   // Kleine Einschatverzögerung
         L     #Temp_SetValueTemp;
         L     "DB751_auxiliaryDriveMetering".HeatexchangerLP[1].Offset_Cooling;
         +R;
         L     #Temp_ND_WT;
         >R;
         =     #Temp_MoreDelta;
   // Kühlen  AUS
         L     "DB613_Komponent_State".HeatexchangerLP[1].PulsTime;
         RND;
         L     #Zeit_abgelaufen;
         <D;
         AN(;
         L     "DB613_Komponent_State".HeatexchangerLP[1].PulsTime;
         RND;
         L     #Regelstrecke;
         >D;
         );
         ON    "DB613_Komponent_State".HeatexchangerLP[1].Switch_Temp_ON_OFF;
         ON    "DB619_State_MPart".Operationmode[1].valid;
         O     "DB823_Error_Metering".Temperature_HeatexchangerLP[1].Sensor_FLT_broken_wire;
         O     #Temp_MoreDelta;
         R     "DB613_Komponent_State".HeatexchangerLP[1].CoolingActive;

   // Valve in FB101 for Heatexchanger in back run
   //      =     "V_Heatexchanger_C1" // stromlos zu

   //-----
   // Check limits temperature 1 Heatexchanger

         CALL  "FC916_PV_Limits"
         ( IN_Tolerance_Test     := "DB619_State_MPart".Operationmode[1].Controllvoltage,
           IN_Reset_Fault        := "DB009_Faults".Faults_Reset_FKT_M1,
           IO_Any_ArrayPV        := "DB608_PV_Metering".HeatexchangerLP[1],
           IO_Fault_Warn_upperL  := "DB823_Error_Metering".Temperature_HeatexchangerLP[1].Warning_limit_plus,
           IO_Fault_Warn_lowerL  := "DB823_Error_Metering".Temperature_HeatexchangerLP[1].Warning_limit_minus,
           IO_Fault_Alarm_upperL := "DB823_Error_Metering".Temperature_HeatexchangerLP[1].Alarm_limit_plus,
           IO_Fault_Alarm_lowerL := "DB823_Error_Metering".Temperature_HeatexchangerLP[1].Alarm_limit_minus,
           IO_New_Fault          := "DB009_Faults".Faultschanging_M1,
           IO_Fault_Level_1      := "DB009_Faults".Faults_FKT_Grp_1_M1,
           IO_Fault_Level_2      := "DB009_Faults".Faults_FKT_Grp_2_M1,
           IO_Fault_Level_3      := "DB009_Faults".Faults_FKT_Grp_3_M1
         );
   //-----
   // State of Switch
         L     0;
         A     "DB613_Komponent_State".HeatexchangerLP[1].CoolingActive;
         A     "DB619_State_MPart".Machine[1].Metering."01";
         A     "DB613_Komponent_State".HeatexchangerLP[1].Switch_Temp_ON_OFF;
         JCN   S1H1;
         L     1;
   S1H1: ON    "DB613_Komponent_State".HeatexchangerLP[1].CoolingActive;
         ON    "DB619_State_MPart".Machine[1].Metering."01";
         A     "DB613_Komponent_State".HeatexchangerLP[1].Switch_Temp_ON_OFF;
         JCN   S2H1;
         L     3;
   S2H1: A     "DB823_Error_Metering".Temperature_HeatexchangerLP[1].Sensor_FLT_broken_wire;
         A     "DB613_Komponent_State".HeatexchangerLP[1].Switch_Temp_ON_OFF;
         JCN   S3H1;
         L     2;
   S3H1: T     "DB613_Komponent_State".HeatexchangerLP[1].State_Temp;
   EHD1: NOP   0;

   // Fault exists
         O     "DB823_Error_Metering".Temperature_HeatexchangerLP[1].Sensor_FLT_broken_wire;
         O     "DB823_Error_Metering".Temperature_HeatexchangerLP[1].Warning_limit_plus;
         O     "DB823_Error_Metering".Temperature_HeatexchangerLP[1].Warning_limit_minus;
         O     "DB823_Error_Metering".Temperature_HeatexchangerLP[1].Alarm_limit_plus;
         O     "DB823_Error_Metering".Temperature_HeatexchangerLP[1].Alarm_limit_minus;
         =     "DB613_Komponent_State".HeatexchangerLP[1].Fault_Exist;
END_REGION

REGION Network 2: There is no connection to the sensor (3)
   //---------------------------------------------
   //  Controller temperature Heatexchanger K2
   //---------------------------------------------
         AN    "DB753_MeteringPump".Pump[2].WithLPHeatExchanger;
         R     "DB823_Error_Metering".Temperature_HeatexchangerLP[2].Sensor_FLT_broken_wire;
         R     "DB823_Error_Metering".Temperature_HeatexchangerLP[2].Warning_limit_plus;
         R     "DB823_Error_Metering".Temperature_HeatexchangerLP[2].Warning_limit_minus;
         R     "DB823_Error_Metering".Temperature_HeatexchangerLP[2].Alarm_limit_plus;
         R     "DB823_Error_Metering".Temperature_HeatexchangerLP[2].Alarm_limit_minus;
         R     "DB613_Komponent_State".HeatexchangerLP[2].Fault_Exist;
         JC    EHD2;
   //-----
         CALL  "FC920_PV_Calc_Act_Value"
         ( IN_Act_Value_read := TRUE,
           IN_Act_Value_ext  := FALSE,
           IN_Ext_Value      := #DINT_dummy,
           IN_Read_Double    := FALSE,
           IN_FLT_Needful    := 1,
           IN_FLT_Reset      := "DB009_Faults".Faults_Reset_FKT_M1,
           IO_Any_ArrayPV    := "DB608_PV_Metering".HeatexchangerLP[2],
           IO_Fault_Sensor   := "DB823_Error_Metering".Temperature_HeatexchangerLP[2].Sensor_FLT_broken_wire,
           IO_New_Fault      := "DB009_Faults".Faultschanging_M1,
           IO_FLT_Level_3    := "DB009_Faults".Faults_FKT_Grp_3_M1
         );
   //
         L     "DB608_PV_Metering".HeatexchangerLP[2].PV_ActV.Value;
         DTR;
         L     10.0;
         /R;
         T     #Temp_ND_WT;
   //
         L     "DB608_PV_Metering".HeatexchangerLP[2].PV_SetV.Value;
         DTR;
         L     10.0;
         /R;
         T     #Temp_SetValueTemp;
   //
         CALL  "FC056_TemPulse2"
         ( Trig              := "Start_Controler1_LP_K2",
           In_Sollwert       := #Temp_SetValueTemp,
           In_Istwert_Tank   := #Temp_ND_WT,
           In_Istwert_Return := #Temp_ND_WT,
           In_Wichtung       := "DB751_auxiliaryDriveMetering".HeatexchangerLP[2].Weighting_Temp,
           In_Regelstrecke   := "DB751_auxiliaryDriveMetering".HeatexchangerLP[2].PLC_Control_Area,
           In_MaxDelta_K     := "DB751_auxiliaryDriveMetering".HeatexchangerLP[2].Max_Temp_Diff_Cooling,
           In_MaxDelta_H     := "DB751_auxiliaryDriveMetering".HeatexchangerLP[2].Max_Temp_Diff_Heating,
           Pulsezeit         := "DB613_Komponent_State".HeatexchangerLP[2].PulsTime,
           Heating           := #Dummy,
           Cooling           := #Temp_Cooling
         );
   //
   //Regelstrecke ms Format
         L     "DB751_auxiliaryDriveMetering".HeatexchangerLP[2].PLC_Control_Area;
         L     1000.0;
         *R;
         RND;
         T     #Regelstrecke;  // Zeitwert für Timer

   // Regelstreckentimer ständig starten

         AN    "Start_Controler1_LP_K2";
         =     "Start_Controler2_LP_K2";

         CALL  TON , "DB61_Temp_ND_WT_MK1_K2"
         ( IN := "Start_Controler2_LP_K2",
           PT := #Regelstrecke,
           Q  := "Start_Controler1_LP_K2",
           ET := #Zeit_abgelaufen
         );

   // Kühlen  EIN
         A     #Temp_Cooling;
         S     "DB613_Komponent_State".HeatexchangerLP[2].CoolingActive;

   //Kleine Einschatverzögerung
         L     #Temp_SetValueTemp;
         L     "DB751_auxiliaryDriveMetering".HeatexchangerLP[2].Offset_Cooling;
         +R;
         L     #Temp_ND_WT;
         >R;
         =     #Temp_MoreDelta;

   // Kühlen  AUS
         L     "DB613_Komponent_State".HeatexchangerLP[2].PulsTime;
         RND;
         L     #Zeit_abgelaufen;
         <D;
         AN(;
         L     "DB613_Komponent_State".HeatexchangerLP[2].PulsTime;
         RND;
         L     #Regelstrecke;
         >D;
         );
         ON    "DB613_Komponent_State".HeatexchangerLP[2].Switch_Temp_ON_OFF;
         ON    "DB619_State_MPart".Operationmode[1].valid;
         O     "DB823_Error_Metering".Temperature_HeatexchangerLP[2].Sensor_FLT_broken_wire;
         O     #Temp_MoreDelta;
         R     "DB613_Komponent_State".HeatexchangerLP[2].CoolingActive;

   // Valve in FB102 for Heatexchanger in back run
   //     =     "V_Heatexchanger_C2" // stromlos zu


   //-----
   // Check limits temperature 2 Heatexchanger

         CALL  "FC916_PV_Limits"
         ( IN_Tolerance_Test     := "DB619_State_MPart".Operationmode[1].Controllvoltage,
           IN_Reset_Fault        := "DB009_Faults".Faults_Reset_FKT_M1,
           IO_Any_ArrayPV        := "DB608_PV_Metering".HeatexchangerLP[2],
           IO_Fault_Warn_upperL  := "DB823_Error_Metering".Temperature_HeatexchangerLP[2].Warning_limit_plus,
           IO_Fault_Warn_lowerL  := "DB823_Error_Metering".Temperature_HeatexchangerLP[2].Warning_limit_minus,
           IO_Fault_Alarm_upperL := "DB823_Error_Metering".Temperature_HeatexchangerLP[2].Alarm_limit_plus,
           IO_Fault_Alarm_lowerL := "DB823_Error_Metering".Temperature_HeatexchangerLP[2].Alarm_limit_minus,
           IO_New_Fault          := "DB009_Faults".Faultschanging_M1,
           IO_Fault_Level_1      := "DB009_Faults".Faults_FKT_Grp_1_M1,
           IO_Fault_Level_2      := "DB009_Faults".Faults_FKT_Grp_2_M1,
           IO_Fault_Level_3      := "DB009_Faults".Faults_FKT_Grp_3_M1
         );
   //-----
   // State of Switch
         L     0;
         A     "DB613_Komponent_State".HeatexchangerLP[2].CoolingActive;
         A     "DB619_State_MPart".Machine[1].Metering."02";
         A     "DB613_Komponent_State".HeatexchangerLP[2].Switch_Temp_ON_OFF;
         JCN   S1H2;
         L     1;
   S1H2: ON    "DB613_Komponent_State".HeatexchangerLP[2].CoolingActive;
         ON    "DB619_State_MPart".Machine[1].Metering."02";
         A     "DB613_Komponent_State".HeatexchangerLP[2].Switch_Temp_ON_OFF;
         JCN   S2H2;
         L     3;
   S2H2: A     "DB823_Error_Metering".Temperature_HeatexchangerLP[2].Sensor_FLT_broken_wire;
         A     "DB613_Komponent_State".HeatexchangerLP[2].Switch_Temp_ON_OFF;
         JCN   S3H2;
         L     2;
   S3H2: T     "DB613_Komponent_State".HeatexchangerLP[2].State_Temp;
   EHD2: NOP   0;

   // Fault exists
         O     "DB823_Error_Metering".Temperature_HeatexchangerLP[2].Sensor_FLT_broken_wire;
         O     "DB823_Error_Metering".Temperature_HeatexchangerLP[2].Warning_limit_plus;
         O     "DB823_Error_Metering".Temperature_HeatexchangerLP[2].Warning_limit_minus;
         O     "DB823_Error_Metering".Temperature_HeatexchangerLP[2].Alarm_limit_plus;
         O     "DB823_Error_Metering".Temperature_HeatexchangerLP[2].Alarm_limit_minus;
         =     "DB613_Komponent_State".HeatexchangerLP[2].Fault_Exist;
END_REGION
END_FUNCTION

FUNCTION "FC071_CleaningPiston" : Void   // FC71, STL
TITLE = Function of cleaning piston mixing head
{ S7_Optimized_Access := 'FALSE' }
AUTHOR : KT242
FAMILY : RS_KK
NAME : CP
VERSION : 1.3
   VAR_INPUT
      IN_WithCP : Bool;   // Signal cleaning piston exists at mixinghead
      IN_Ana_CP_State : Byte;   // State of analog cleaning piston
      IN_SWUEnabled : Bool;   // Switch over unit for this mixing head is enabled
      IN_ButtonCPForward : Bool;   // Button cleaning piston manually forward
      IN_ButtonCPback : Bool;   // Button cleaning piston manually back
      IN_CPForwardFromExternal : Bool;   // External signal (e.g. from robot) to move the CP forward
      IN_CPAfterShot : Bool;   // Signal cleaning piston has to move after the shot
      IN_PartshotDisabled : Bool;   // Partshot disabled -> like service shot
      IN_Blowing_OUT : Bool;   // Blowing out after Shot
      IN_CPProxSwitch : Bool;   // Proximity switch cleaning piston is back (rest position)
      IN_SWUActive : Bool;   // Only this switch over unit is activated
      IN_HydraulicOk : Bool;   // Hydraulic ok
      IN_ResetFaults : Bool;   // Signal to reset error bits
      IN_ControlVoltage : Bool;   // Control Voltage is on
      IN_OperatingModeValid : Bool;   // Valid operating mode is activated
      IN_OperatingModeWithFoam : Bool;   // Machine is not in service mode (this is a condition for cleaning)
      IN_OperatingModeTestValv : Bool;   // Machine is in mode test with test valves (no cleaning necessary)
      IN_Lamptest : Bool;   // Lamptest selected
      IN_ShotEnd : Bool;   // Ramp shot finished
      IN_FaultLevel_1 : Bool;   // Fault level 1 on machine
      IN_PressurizeTimeRunning : Bool;   // Time for building up pressure and flow values is active
      IN_ShotActive : Bool;   // Shot is active
      IN_CycleRunning : Bool;   // Shotcycle is active
      IN_RmpCtrlChangeTimeEnd : Bool;   // Recirculation between shots finished
      IN_StandbyTimeRunning : Bool;   // Recirculation after shot acvtiv
      IN_RmpCycleEnd : Bool;   // Foaming cycle finished
      IN_CPTimer : Timer;   // Timer for CP-funkctions
      IN_TMCheckHomePos : Timer;   // Timer to suppress fault homepos when module begins regulation
      Values : "UDT771_CleaningPiston";
   END_VAR
   VAR_IN_OUT
      OUT_ValveCPForward : Bool;   // Valve to move the CP forward
      OUT_LampCPBack : Bool;   // Lamp to display that the CP is back
      IO_CPIsOk : Bool;   // CP is ok -> enables shot
      IO_ReqHydrForCleaning : Bool;   // Request hydraulic pressure for cleaning stroke
      IO_Status : ANY;   // Status flags for CP
      IO_Fault : ANY;
      IO_NewFault : Bool;
      IO_FaultLevel_1 : Bool;
      IO_FaultLevel_2 : Bool;
      IO_FaultLevel_3 : Bool;
   END_VAR
   VAR_TEMP
      Temp_IO_Status : "UDT071_CPiston_State";
      TEMP_IO_Fault : "UDT1871_FLT_CPiston";
      ERROR_CODE : Int;   // Error state of systemfunction "BLKMOV" Blockmove
      Anypointer1 : ANY;   // Pointer to copy thr array "IO_Status" and "Temp_IO_Status"
      Anypointer2 : ANY;   // Pointer to copy thr array "IO_Status" and "Temp_IO_Status"
      InterruptCleaningStroke : Bool;   // Flag of interrupt cleaning cycle
      StartCleaningStroke : Bool;   // Flag cleaning cycle started
      ShotFinished : Bool;   // Flag activate cleaning piston after part shot
      TempAnaCPBack : Bool;   // Analog controlled leaning piston is back
      WrongType : Bool;   // Wrong Mixing Head Type
   END_VAR
BEGIN

REGION Network 1: Saved data integration
         LAR1;
         L;
         LAR2;
   //
         L     16#1002;  // Bytes
         T     W[AR1, P#0.0];
         L     W[AR2, P#2.0];  // Amount of bytes
         T     W[AR1, P#2.0];
         L     W[AR2, P#4.0];  // Block no,
         T     W[AR1, P#4.0];
         L     D[AR2, P#6.0];  // Startadress of datas
         T     D[AR1, P#6.0];
   //
         CALL  BLKMOV
         ( SRCBLK  := #Anypointer1,
           RET_VAL := #ERROR_CODE,
           DSTBLK  := #Temp_IO_Status
         );
   //
         LAR1;
         L;
         LAR2;
   //
         L     16#1002;  // Bytes
         T     W[AR1, P#0.0];
         L     W[AR2, P#2.0];  // Amount of bytes
         T     W[AR1, P#2.0];
         L     W[AR2, P#4.0];  // Block no,
         T     W[AR1, P#4.0];
         L     D[AR2, P#6.0];  // Startadress of datas
         T     D[AR1, P#6.0];
   //
         CALL  BLKMOV
         ( SRCBLK  := #Anypointer2,
           RET_VAL := #ERROR_CODE,
           DSTBLK  := #TEMP_IO_Fault
         );
   //
         A(;
         L     #IN_Ana_CP_State;
         AW    16#0080;
         A     <>0;
         );
         A(;
         O     #Values.ContrCleaningPiston;
         O     #Values.StepCleaningPiston;
         );
         =     #TempAnaCPBack;
END_REGION

REGION Network 2: Cleaning stroke forward
         AN    #IN_WithCP;
         R     #Values.Spare_19;

         ON    #IN_WithCP;
         ON    #Values.Spare_19;
         R     #Temp_IO_Status.Switch_CP_Forward;

         NOT;
         CLR;
         =     #WrongType;
         A     #WrongType;
         JC    STG;
END_REGION

REGION Network 3: CP existing or not?
         O     #IN_CPProxSwitch;
         O     #TempAnaCPBack;
         AN    #TEMP_IO_Fault.IPS_defect;
         ON    #IN_WithCP;
         A     #IN_SWUActive;
         =     #Temp_IO_Status.CP_is_OK;
         S     #IO_CPIsOk;
   //
         A     #Temp_IO_Status.CP_is_OK;
         FN    #Temp_IO_Status.Edge_CP_nOK;
         R     #IO_CPIsOk;
   //
         A     #IN_SWUEnabled;
         A     #IN_WithCP;
         JC    STG;
   //
         SET;
         R     #Temp_IO_Status.MH_was_open;
         R     #Temp_IO_Status.Cleaning_runs;
         R     #Temp_IO_Status.CleaningFromEPrunning;
         R     #Temp_IO_Status.CleanAfterShotSelected;
         R     #Temp_IO_Status.Stop_Cleaning;
         R     #Temp_IO_Status.CP_valve_selected;
         R     #Temp_IO_Status.CP_Moved_Manual;
         R     #Temp_IO_Status.FaultExists;
         R     #TEMP_IO_Fault.Forward_to_slow;
         R     #TEMP_IO_Fault.Back_to_slow;
         R     #TEMP_IO_Fault.IPS_defect;
         R     #TEMP_IO_Fault.Lost_IPS_position;
         L     0;
         T     #Temp_IO_Status.Stepnumber;
   //
         JU    LAMP;
END_REGION

REGION Network 4: Error handling
   STG:  NOP   0;
   // Reset faults
         A     #IN_ResetFaults;
         R     #TEMP_IO_Fault.Lost_IPS_position;
         R     #TEMP_IO_Fault.IPS_defect;
         R     #TEMP_IO_Fault.Forward_to_slow;
         R     #TEMP_IO_Fault.Back_to_slow;
         R     #TEMP_IO_Fault.Leaves_HomePos;
   //
         A     #WrongType;
         JC    err;

   // Fault No.1: Cleaning piston leaves the backward position during shot
         L     2#0000_0000_0000_0100;
         L     #IN_Ana_CP_State;
         AW;
         L     0;
         >D;
         A(;
         O     #Values.ContrCleaningPiston;
         O     #Values.StepCleaningPiston;
         );
         O;
         A     #IN_SWUActive;
         A     #IN_ShotActive;
         AN(;
         O     #Values.ContrCleaningPiston;
         O     #Values.StepCleaningPiston;
         );
         AN    #IN_CPProxSwitch;
         AN    #TEMP_IO_Fault.Lost_IPS_position;
         S     #TEMP_IO_Fault.Lost_IPS_position;
         S     #IO_NewFault;
   //
   // Fault No.2: Priximity switch cleaning piston back is broken
         AN    #IN_CPProxSwitch;
         A     #IN_HydraulicOk;
         AN    #TEMP_IO_Fault.Back_to_slow;
         AN    #Temp_IO_Status.Cleaning_runs;
         AN(;
         O     #Values.ContrCleaningPiston;
         O     #Values.StepCleaningPiston;
         );
         AN    #TEMP_IO_Fault.Lost_IPS_position;
         AN    #TEMP_IO_Fault.IPS_defect;
         S     #TEMP_IO_Fault.IPS_defect;
         S     #IO_NewFault;
   //
   // Fault No. 3: Movement forward of analog cleaning piston too slow
         L     2#0000_0000_0000_0001;
         L     #IN_Ana_CP_State;
         AW;
         L     0;
         >D;
         A(;
         O     #Values.ContrCleaningPiston;
         O     #Values.StepCleaningPiston;
         );
         AN    #TEMP_IO_Fault.Forward_to_slow;
         S     #TEMP_IO_Fault.Forward_to_slow;
         S     #IO_NewFault;
   // Fault No. 3: Movement forward of cleaning piston too slow is build later
   //

   // Fault No. 4: Movement back of analog cleaning piston too slow
         L     2#0000_0000_0000_0010;
         L     #IN_Ana_CP_State;
         AW;
         L     0;
         >D;
         A(;
         O     #Values.ContrCleaningPiston;
         O     #Values.StepCleaningPiston;
         );
         AN    #TEMP_IO_Fault.Back_to_slow;
         S     #TEMP_IO_Fault.Back_to_slow;
         S     #IO_NewFault;
   // Fault No. 4: Movement back of cleaning piston too slow is build later
   //
   // Fault No. 14: Cleaning piston is leaving home position
   //
         A     #IN_HydraulicOk;
         L     S5T#500MS;
         SD    #IN_TMCheckHomePos;
         A(;
         L     2#0000_0000_0010_0000;
         L     #IN_Ana_CP_State;
         AW;
         L     0;
         >D;
         );
         A(;
         O     #Values.ContrCleaningPiston;
         O     #Values.StepCleaningPiston;
         );
         A     #IN_TMCheckHomePos;
         AN    #TEMP_IO_Fault.Leaves_HomePos;
         S     #TEMP_IO_Fault.Leaves_HomePos;
         S     #IO_NewFault;
END_REGION

REGION Network 5: Error handling
   err:  NOP   0;
         O     #TEMP_IO_Fault.Forward_to_slow;
         O     #TEMP_IO_Fault.Back_to_slow;
         O     #TEMP_IO_Fault.IPS_defect;
         O     #TEMP_IO_Fault.Lost_IPS_position;
         O     #TEMP_IO_Fault.Leaves_HomePos;
         =     #Temp_IO_Status.FaultLevel_1;
         =     #Temp_IO_Status.FaultExists;
         S     #IO_FaultLevel_1;

         CLR;
         =     #Temp_IO_Status.FaultLevel_2;
         S     #IO_FaultLevel_2;

         CLR;
         =     #Temp_IO_Status.FaultLevel_3;
         S     #IO_FaultLevel_3;

         A     #WrongType;
         JC    LAMP;
END_REGION

REGION Network 6: Cleaning necessary or not
   // Step 1: Detect if the mixinghead was open.
   //         The signal is built newly for each partshot and only if the mixinghead
   //         was really opened a cleaning stroke is carried out
   //         -> "Temp_IO_Status.MH_was_open"
   //         It is reset when:
   //         - the switching unit is deselected
   //         - a new shot is started (no matter on wich mixinghead)
   //         - the shot cycle is finished
   //         - the cleaning stroke was done
   //         - the operating mode is deselected
   // 
   // Step 2: If for this shot a cleaning stroke was selected or after fault group 1
   //         the cleaning piston moves forward.
   //         -> "Temp_IO_Status.Cleaning_a_Shot_selected"
   //         The bit is reset if:
   //         - the switching unit is deselected
   //         - the cleaning stroke was done 
   //         - the operating mode is deselected
         A     #IN_ShotActive;
         A     #IN_OperatingModeWithFoam;
         AN    #IN_PartshotDisabled;
         AN    #IN_OperatingModeTestValv;
         A     #IN_SWUActive;
         S     #Temp_IO_Status.MH_was_open;
   //
         A     #IN_CPAfterShot;
         A     #IN_ShotEnd;
         O     #IN_FaultLevel_1;
         ON    #IN_ControlVoltage;
         A     #Temp_IO_Status.MH_was_open;
         S     #Temp_IO_Status.CleanAfterShotSelected;
   //
         O     #Temp_IO_Status.CleanAfterShotSelected;
         O     #IN_RmpCtrlChangeTimeEnd;
         O     #Temp_IO_Status.Stop_Cleaning;
         ON    #IN_OperatingModeValid;
         R     #Temp_IO_Status.MH_was_open;
   //
END_REGION

REGION Network 7: Interrupt cleaning stroke
   // A cleaning cycle is interrupted in the following cases:
   //            - Button cleaning piston back is used without acting the butten
   //              cleaning piston forward at the same time  (LFI) 
   //            - The robot resets the signal cleaning piston forward
   //            - a new shot is being started on this mixinghead
   // 
   // If a cleaning stroke should be interrupted, the step counter for the cleaning
   // cycle is set to 6 (reset output for valve CP forward)
         A(;
         O     #IN_PressurizeTimeRunning;
         O     #IN_RmpCtrlChangeTimeEnd;
         A     #IN_SWUActive;
         O;
         A     #Temp_IO_Status.CleaningFromEPrunning;
         AN    #IN_CPForwardFromExternal;
         O;
         A     #IN_ButtonCPback;
         );
         A     #Temp_IO_Status.Cleaning_runs;
         AN    #Temp_IO_Status.Stop_Cleaning;
         S     #Temp_IO_Status.Stop_Cleaning;
         =     #InterruptCleaningStroke;
   //
         AN    #InterruptCleaningStroke;
         JC    CONT;
   //
         L     6;
         T     #Temp_IO_Status.Stepnumber;
   //
   CONT: A     #IN_CPForwardFromExternal;
         =     #Temp_IO_Status.CleaningFromEPrunning;
END_REGION

REGION Network 8: Start cleaning stroke
   //  1. Block:
   //
         A(;
   // A.:
         O     #IN_ButtonCPForward;
         O     #Temp_IO_Status.Switch_CP_Forward;
         AN    #IN_ButtonCPback;
         O     #Temp_IO_Status.CleaningFromEPrunning;
         A(;
         ON    #IN_CycleRunning;
         O     #IN_StandbyTimeRunning;
         ON    #IN_SWUActive;
         );
   // B.:
         O(;
         A     #IN_ShotEnd;
         A     #Temp_IO_Status.CleanAfterShotSelected;
         );
         );
         A     #IN_HydraulicOk;
   //  2. Block:
   //
         O(;
         ON    #IN_ControlVoltage;
         O     #IN_FaultLevel_1;
         A     #Temp_IO_Status.CleanAfterShotSelected;
         );
   // für alle:
         AN    #Temp_IO_Status.Stop_Cleaning;
         AN    #Temp_IO_Status.Cleaning_runs;
         S     #Temp_IO_Status.Cleaning_runs;
         =     #StartCleaningStroke;
   //
         AN    #StartCleaningStroke;
         JC    STEP;
   //
         A     #IN_ButtonCPForward;
         S     #Temp_IO_Status.CP_Moved_Manual;
         L     1;
         T     #Temp_IO_Status.Stepnumber;
   STEP: NOP   0;
END_REGION

REGION Network 9: organize steps of cleaning stroke
         L     #Temp_IO_Status.Stepnumber;
         JL    DEL;  // if step number > 7 or
         JU    DEL;  // 0: delete
         JU    ST1;  // 1: check if waiting time back needs to be started
         JU    ST2;  // 2: start waiting time back
         JU    ST3;  // 3: actuate the valve
         JU    ST4;  // 4: monitor movement time forward
         JU    ST5;  // 5: start wait time in front
         JU    ST6;  // 6: switch off valve for CP
         JU    ST7;  // 7: monitor movement back
   //
   DEL:  CLR;  // delete status informations
         =     #Temp_IO_Status.CP_valve_selected;
         =     #Temp_IO_Status.Cleaning_runs;
         =     #Temp_IO_Status.Stop_Cleaning;
         CLR;
         SP    #IN_CPTimer;
         JU    LAMP;
END_REGION

REGION Network 10: check: wait time back necessary
   ST1:  SET;
         R     #Temp_IO_Status.Stop_Cleaning;
   //
         A     #Temp_IO_Status.CleanAfterShotSelected;
         JCN   ST1E;
         L     2;  // start waiting time back (if automatic cleaning stroke)
         T     #Temp_IO_Status.Stepnumber;
         JU    LAMP;
   //
   ST1E: L     3;  // start cleaning directly (in other cases)
         T     #Temp_IO_Status.Stepnumber;
         JU    LAMP;
END_REGION

REGION Network 11: start waiting time back
   // The waitint time back normally is 0.2 seconds
   ST2:  AN    #IN_Blowing_OUT;
         L     #Values.RestTimeBack;
         SD    #IN_CPTimer;
         AN    #IN_CPTimer;
         JC    LAMP;
   //
         L     3;
         T     #Temp_IO_Status.Stepnumber;
         CLR;
         SP    #IN_CPTimer;
         JU    LAMP;
END_REGION

REGION Network 12: Actuate the valve
   ST3:  SET;
         S     #Temp_IO_Status.CP_valve_selected;
         S     #IO_ReqHydrForCleaning;
         L     4;
         T     #Temp_IO_Status.Stepnumber;
         JU    LAMP;
END_REGION

REGION Network 13: Monitor movement time forward
   // the monitoring time is fix on 2 seconds
   ST4:  O     #IN_CPProxSwitch;  // next step when prximity switch is off
         O     #TempAnaCPBack;
         JC    LZVW;
   //
         L     5;
         T     #Temp_IO_Status.Stepnumber;
         CLR;
         SP    #IN_CPTimer;
         JU    LAMP;
   //
   LZVW: L     S5T#2S;
         SD    #IN_CPTimer;
         A     #IN_CPTimer;
         JCN   LAMP;
   //
   // Fault No.3: movement forward too slow
   //
         R     #Temp_IO_Status.CleanAfterShotSelected;
         AN    #TEMP_IO_Fault.Forward_to_slow;
         S     #TEMP_IO_Fault.Forward_to_slow;
         S     #IO_NewFault;
         L     0;
         T     #Temp_IO_Status.Stepnumber;
         JU    LAMP;
END_REGION

REGION Network 14: Wait time in fromt
   //-----
   ST5:  SET;
         R     #Temp_IO_Status.CleanAfterShotSelected;
   //-----
         A     #Temp_IO_Status.CP_Moved_Manual;
         L     #Values.RestTimeFrontManual;
         JC    TimeCPForward;
         L     #Values.RestTimeFront;
   //-----
   TimeCPForward:NOP   0;
         SET;
         SD    #IN_CPTimer;
   //-----
         A     #IN_CPTimer;
         AN    #IN_ButtonCPForward;
         AN    #Temp_IO_Status.Switch_CP_Forward;
         AN    #Temp_IO_Status.CleaningFromEPrunning;
         JCN   LAMP;
   //-----
         L     6;
         T     #Temp_IO_Status.Stepnumber;
         CLR;
         SP    #IN_CPTimer;
         JU    LAMP;
   //-----
END_REGION

REGION Network 15: switch off the valve
   ST6:  SET;
         S     #Temp_IO_Status.Stop_Cleaning;
         R     #Temp_IO_Status.CP_valve_selected;
         R     #Temp_IO_Status.CP_Moved_Manual;
         S     #IO_ReqHydrForCleaning;
         L     7;
         T     #Temp_IO_Status.Stepnumber;
         CLR;
         SP    #IN_CPTimer;
         JU    LAMP;
END_REGION

REGION Network 16: monitoring movement back
   ST7:  CLR;
         AN    #IN_CPProxSwitch;
         AN    #TempAnaCPBack;
         AN    #TEMP_IO_Fault.Back_to_slow;
         JC    ST7E;
   //
         L     0;
         T     #Temp_IO_Status.Stepnumber;
         SET;
         R     #Temp_IO_Status.Cleaning_runs;
         CLR;
         SP    #IN_CPTimer;
         JU    LAMP;
   //
   ST7E: L     S5T#5S;
         SD    #IN_CPTimer;
         A     #IN_CPTimer;
   //
   // Fault No.4: movement back too slow
   //
         AN    #TEMP_IO_Fault.Back_to_slow;
         S     #TEMP_IO_Fault.Back_to_slow;
         S     #IO_NewFault;
         JU    LAMP;
END_REGION

REGION Network 17: actuate valve and lamp
   LAMP: O     #IN_CPProxSwitch;
         O     #TempAnaCPBack;
         O     #IN_Lamptest;
         AN    #WrongType;
         =     #OUT_LampCPBack;
   //
         A     #Temp_IO_Status.CP_valve_selected;
         AN    #WrongType;
         =     #OUT_ValveCPForward;
END_REGION

REGION Network 18: State of drive: 1-> Selected and ON; 2->Selected but not ON; 3->Not Selected but ON; 4-> Faulty
   //-----
         L     0;
         O     #IN_CPProxSwitch;
         O     #TempAnaCPBack;
         A     #Temp_IO_Status.CP_valve_selected;
         L     1;
         JU    tran;
   //-----
         AN    #OUT_LampCPBack;
         A     #Temp_IO_Status.CP_valve_selected;
         L     2;
         JU    tran;
   //-----
         CLR;
         L     3;
         JU    tran;
   //-----
         O     #Temp_IO_Status.FaultLevel_1;
         O     #Temp_IO_Status.FaultLevel_2;
         O     #Temp_IO_Status.FaultLevel_3;
         L     4;
         JU    tran;
   //-----
   tran: T     #Temp_IO_Status.State_CP;
   //-----
END_REGION

REGION Network 19: Save data
         CALL  BLKMOV
         ( SRCBLK  := #Temp_IO_Status,
           RET_VAL := #ERROR_CODE,
           DSTBLK  := #Anypointer1
         );
   //
         CALL  BLKMOV
         ( SRCBLK  := #TEMP_IO_Fault,
           RET_VAL := #ERROR_CODE,
           DSTBLK  := #Anypointer2
         );
   //
END_REGION
END_FUNCTION

FUNCTION "FC081_FaultsGen" : Void   // FC81, STL
TITLE = General faults of a pouring machine
{ S7_Optimized_Access := 'FALSE' }
AUTHOR : KT242
FAMILY : RS_KK
NAME : Fault_M1
VERSION : 1.1
   VAR_INPUT
      IN_Erster_SPS_Zyklus : Bool;   // Impulssignal Neusstart der Steuerung zum ablöschen der Störungen
   END_VAR
   VAR_TEMP
      ERROR_CODE : Int;   // Error state of systemfunction "BLKMOV" Blockmove
      Null : Word;
      Temp_MinShotTime : Time;
      Temp_MinShotTime_INT : DInt;
   END_VAR
BEGIN

REGION Network 1: Reset general faults
         A     "DB009_Faults".Faults_Reset_FKT_M1;
         JCN   nres;

         L     0;
         T     #Null;

         CALL  FILL
         ( BVAL    := #Null,
           RET_VAL := #ERROR_CODE,
           BLK     := "DB820_Error_general".Machine[1]
         );

         CALL  FILL
         ( BVAL    := #Null,
           RET_VAL := #ERROR_CODE,
           BLK     := "DB820_Error_general".Machine[2]
         );

   nres: NOP   0;
END_REGION

REGION Network 2: Fault level 1

   // Data lost after erasing PLC  -- DB810.DBX 64.0
   //    UN    DB11.DBX  417.0
   //    S     "DB820_Error_general".Machine[1].Data_lost_after_erasing
   //    U     "DB820_Error_general".Machine[1].Data_lost_after_erasing
   //    FP    #IO_Fault.Data_lost_after_erasing
   //    S     "DB009_Faults".Faultschanging_M1

   // Operationmode cylinder service not permitted  DB810.DBX 64.6
   //    O     "S_BA_Automatik"
   //    O     "DB619_State_MPart".Recirculation_Ma[1].Reduced
   //    O     "DB619_State_MPart".Recirculation_Ma[1].Highpressure
   //    O     "DB619_State_MPart".Recirculation_Ma[1].Pausetime
   //    O     "DB619_State_MPart".Recirculation_Ma[1].Lowpressure
   //    O     "DB619_State_MPart".Recirculation_Ma[1].Weekendswitching
   //    U     "DB619_State_MPart".CylinderManager_Ma[1].Cylinderservice
   //    U     "DB619_State_MPart".CylinderManager_Ma[1].Block_is_active
   //    UN    "DB820_Error_general".Machine[1].CylinderServiceNotPermit
   //    S     "DB820_Error_general".Machine[1].CylinderServiceNotPermit
   //    S     "DB009_Faults".Faultschanging_M1

   // Wrong mixinghead no machine 1 -- DB810.DBX 65.3
         O(;
         A(;
         L     1;
         L     "DB619_State_MPart".ShotMa[1].ShotData.MH_No;
         <>I;
         );
         A(;
         O     "DB110_Interf_Program_M1".Status_IF[1].IF_is_on_1_Position;
   //      O     "DB110_Interf_Program_M1".Status_IF[2].IF_is_on_1_Position
   //      O     "DB110_Interf_Program_M1".Status_IF[3].IF_is_on_1_Position
   //      O     "DB110_Interf_Program_M1".Status_IF[4].IF_is_on_1_Position
   //      O     "DB110_Interf_Program_M1".Status_IF[5].IF_is_on_1_Position
         );
         );
   //-
         O(;
         A(;
         L     1;
         L     "DB619_State_MPart".ShotMa[1].ShotData.MH_No;
         <>I;
         );
         A     "DB110_Interf_Program_M1".Status_IF[2].IF_is_on_1_Position;
         );
   //-
         O(;
         A(;
         L     1;
         L     "DB619_State_MPart".ShotMa[1].ShotData.MH_No;
         <>I;
         );
         A     "DB110_Interf_Program_M1".Status_IF[3].IF_is_on_1_Position;
         );
   //-
         O(;
         A(;
         L     1;
         L     "DB619_State_MPart".ShotMa[1].ShotData.MH_No;
         <>I;
         );
         A     "DB110_Interf_Program_M1".Status_IF[4].IF_is_on_1_Position;
         );
   //-
         O(;
         A(;
         L     1;
         L     "DB619_State_MPart".ShotMa[1].ShotData.MH_No;
         <>I;
         );
         A     "DB110_Interf_Program_M1".Status_IF[5].IF_is_on_1_Position;
         );
   //-
         O(;
         A(;
         L     6;
         L     "DB619_State_MPart".ShotMa[1].ShotData.MH_No;
         <>I;
         );
         A     "DB110_Interf_Program_M1".Status_IF[6].IF_is_on_1_Position;
         );
   //-
         O(;
         A(;
         L     7;
         L     "DB619_State_MPart".ShotMa[1].ShotData.MH_No;
         <>I;
         );
         A     "DB110_Interf_Program_M1".Status_IF[7].IF_is_on_1_Position;
         );
   //-
         O(;
         A(;
         L     8;
         L     "DB619_State_MPart".ShotMa[1].ShotData.MH_No;
         <>I;
         );
         A     "DB110_Interf_Program_M1".Status_IF[8].IF_is_on_1_Position;
         );
   //-
         O(;
         A(;
         L     9;
         L     "DB619_State_MPart".ShotMa[1].ShotData.MH_No;
         <>I;
         );
         A     "DB110_Interf_Program_M1".Status_IF[9].IF_is_on_1_Position;
         );
   //-
         O(;
         A(;
         L     10;
         L     "DB619_State_MPart".ShotMa[1].ShotData.MH_No;
         <>I;
         );
         A     "DB110_Interf_Program_M1".Status_IF[10].IF_is_on_1_Position;
         );
   //-
         AN(;
         L     "DB619_State_MPart".ShotMa[1].ShotData.MH_No;
         L     0;
         ==I;
         );
   //-
         A(;
         O     "DB619_State_MPart".Cycle[1].PressurizeTimeRuns;
         O     "DB619_State_MPart".Cycle[1].CtrlChangeTimeRuns;
         );
         AN    "DB619_State_MPart".Operationmode[1].Test;
         AN    "DB820_Error_general".Machine[1].WrongMH_No;
         S     "DB820_Error_general".Machine[1].WrongMH_No;
         S     "DB009_Faults".Faultschanging_M1;

   // Wrong mixinghead no machine 2 -- DB810.DBX 83.3
   //    O(
   //    U(
   //    L     1
   //    L     "DB619_State_MPart".ToolMa[2].ToolNo
   //    <>I
   //    )
   //    U     "DB112_Interf_Program_M2".Status_IF01.IF_is_on_1_Position
   //    )
   //    O(
   //    U(
   //    L     2
   //    L     "DB619_State_MPart".ToolMa[2].ToolNo
   //    <>I
   //    )
   //    U     "DB112_Interf_Program_M2".Status_IF02.IF_is_on_1_Position
   //    )
   //    UN    "DB619_State_MPart".Operationmode_Ma[2].Test
   //    UN    "DB820_Error_general".Machine[2].WrongMH_No
   //    S     "DB820_Error_general".Machine[2].WrongMH_No
   //    S     "DB009_Faults".Faultschanging_M2


   // Alarm Pentan -- DB810.DBX 76.5
   //    UN    "K_AlarmN2_K1"
   //    UN    "DB820_Error_general".Machine[1].FLT_alarm_pentan
   //    S     "DB820_Error_general".Machine[1].FLT_alarm_pentan
   //    S     "DB009_Faults".Faultschanging_M1

   // Fault level 1 from PUC
         A     "DB009_Faults".FaultPC_Level_1;
         AN    "DB820_Error_general".Machine[1].FaultPC_Level_1;
         S     "DB820_Error_general".Machine[1].FaultPC_Level_1;
         S     "DB009_Faults".Faultschanging_M1;

   // Fault level 1 from PUC
   //    U     "DB009_Faults".FaultPC_Level_1
   //    UN    "DB820_Error_general".Machine[2].FaultPC_Level_1
   //    S     "DB820_Error_general".Machine[2].FaultPC_Level_1
   //    S     "DB009_Faults".Faultschanging_M2

   // Buffer shot result full -- DB810.DBX 77.4
   //    U     "DB619_State_MPart".BufferShotResultSignal.FaultBufferFull
   //    UN    "DB820_Error_general".Machine[1].BufferShotDataFull
   //    S     "DB820_Error_general".Machine[1].BufferShotDataFull
   //    S     "DB009_Faults".Faultschanging_M1

   // Buffer shot result full -- DB810.DBX 77.4
   //    U     "DB619_State_MPart".BufferShotResultSignal.FaultBufferFull
   //    UN    "DB820_Error_general".Machine[2].BufferShotDataFull
   //    S     "DB820_Error_general".Machine[2].BufferShotDataFull
   //    S     "DB009_Faults".Faultschanging_M2

   // Foaming time too short-- DB810.dbx78.0

         L     "DB700_Machine".Machine[1].Min_ShotTime;

         CALL  T_CONV
         ( IN  := "DB700_Machine".Machine[1].Min_ShotTime,
           OUT := #Temp_MinShotTime
         );
   //-
         L     #Temp_MinShotTime;
         T     #Temp_MinShotTime_INT;
   //-
         L     "DB606_PV_Machine".Machine[1].ShotTime.PV_SetV.Value;
         L     #Temp_MinShotTime_INT;
         <D;
         A     "DB619_State_MPart".Cycle[1].Shotrelease;
         AN    "DB820_Error_general".Machine[1].ShotTimeTooShort;
         S     "DB820_Error_general".Machine[1].ShotTimeTooShort;
         S     "DB009_Faults".Faultschanging_M1;

   // Foaming time too short-- DB810.dbx78.0
   //    L     "DB606_PV_Machine".Machine[2].ShotTime.PV_SetV.Set_Value
   //    L     250
   //    <D
   //    U     "DB619_State_MPart".Cycle_Ma[2].Shotrelease
   //    UN    "DB820_Error_general".Machine[2].ShotTimeTooShort
   //    S     "DB820_Error_general".Machine[2].ShotTimeTooShort
   //    S     "DB009_Faults".Faultschanging_M2


   // Set fault level 1 machine 1 and 2
         O     "DB820_Error_general".Machine[1].CylinderServiceNotPermit;
   //    O     "DB820_Error_general".Machine[1].BufferShotDataFull
   //    O     "DB820_Error_general".Machine[1].FaultPC_Level_1
   //    O     "DB820_Error_general".Machine[1].Data_lost_after_erasing
         O     "DB820_Error_general".Machine[1].FLT_alarm_pentan;
         O     "DB820_Error_general".Machine[1].WrongMH_No;
         O     "DB820_Error_general".Machine[1].ShotTimeTooShort;
         S     "DB009_Faults".Faults_FKT_Grp_1_M1;

   //    O     "DB820_Error_general".Machine[2].CylinderServiceNotPermit
   //    O     "DB820_Error_general".Machine[2].BufferShotDataFull
   //    O     "DB820_Error_general".Machine[2].FaultPC_Level_1
   //    O     "DB820_Error_general".Machine[2].Data_lost_after_erasing
         O     "DB820_Error_general".Machine[2].FLT_alarm_pentan;
         O     "DB820_Error_general".Machine[2].WrongMH_No;
         O     "DB820_Error_general".Machine[2].ShotTimeTooShort;
         S     "DB009_Faults".Faults_FKT_Grp_1_M2;
END_REGION

REGION Network 3: Fault level 2
   // Störung Gruppe 2 von PC
   //    U     "DB009_Faults".FaultPC_Level_2
   //    UN    "DB820_Error_general".Machine[1].FaultPC_Level_2
   //    S     "DB820_Error_general".Machine[1].FaultPC_Level_2
   //    S     "DB009_Faults".Faultschanging_M1

   //    U     "DB009_Faults".FaultPC_Level_2
   //    UN    "DB820_Error_general".Machine[2].FaultPC_Level_2
   //    S     "DB820_Error_general".Machine[2].FaultPC_Level_2
   //    S     "DB009_Faults".Faultschanging_M2

   //    O     "DB820_Error_general".Machine[1].FaultPC_Level_2
   //    S     "DB009_Faults".Faults_FKT_Grp_2_M1

   //    O     "DB820_Error_general".Machine[2].FaultPC_Level_2
   //    S     "DB009_Faults".Faults_FKT_Grp_2_M2

   // Fault Pneumatik Überwachung
         AN    "P_air";
         AN    "DB820_Error_general".Machine[1].Pneumatik_1;
         CLR;
         S     "DB820_Error_general".Machine[1].Pneumatik_1;
         S     "DB009_Faults".Faultschanging_M1;

   // Fault Pneumatik sanfte Überwachung
         AN    "P_air_2";
         AN    "DB820_Error_general".Machine[1].Pneumatik_2;
         CLR;
         S     "DB820_Error_general".Machine[1].Pneumatik_2;
         S     "DB009_Faults".Faultschanging_M1;

         O     "DB820_Error_general".Machine[1].Pneumatik_1;
         O     "DB820_Error_general".Machine[1].Pneumatik_2;
         S     "DB009_Faults".Faults_FKT_Grp_2_M1;
END_REGION

REGION Network 4: Fault level 3
   // Schnittstelle zum Rechner ist gestört  -- DB810.DBX 76.2
   //    UN    "Merker_Schnittstelle_ok"
   //    UN    "DB820_Error_general".Machine[1].Interface_PC
   //    S     "DB820_Error_general".Machine[1].Interface_PC
   //    S     "DB009_Faults".Faultschanging_M1

   // Pufferbatterie SPS leer  -- DB810.DBX 76.3
   //    U     "Flag_Pufferbatterie"
   //    UN    "DB820_Error_general".Machine[1].BufferBattery
   //    S     "DB820_Error_general".Machine[1].BufferBattery
   //    S     "DB009_Faults".Faultschanging_M1

   // Faulte Fuse machine 1 -- DB810.DBX 64.1
         AN    "F_Fuse_Machine";
         AN    "DB820_Error_general".Machine[1].Fuse_broken;
         S     "DB820_Error_general".Machine[1].Fuse_broken;
         S     "DB009_Faults".Faultschanging_M1;

   // Faulte Fuse machine 2 --
   //    UN    "F_Fuse_Machine_M2"
   //    UN    "DB820_Error_general".Machine[2].Fuse_broken
   //    S     "DB820_Error_general".Machine[2].Fuse_broken
   //    S     "DB009_Faults".Faultschanging_M2

   // Faulte Fuse mixinghead machine 1
         AN    "F_Fuse_MH";
         AN    "DB820_Error_general".Machine[1].Fuse_brocken_Mixinghead;
         S     "DB820_Error_general".Machine[1].Fuse_brocken_Mixinghead;
         S     "DB009_Faults".Faultschanging_M1;

   // Faulte Fuse mixinghead machine 2
   //    UN    "F_Fuse_MH_M2"
   //    UN    "DB820_Error_general".Machine[2].Fuse_brocken_Mixinghead
   //    S     "DB820_Error_general".Machine[2].Fuse_brocken_Mixinghead
   //    S     "DB009_Faults".Faultschanging_M2

   // Fault air dryer -- DB810.DBX 64.4
         AN    "F_Airdryer";
         AN    "DB820_Error_general".Machine[1].Air_dryer;
         S     "DB820_Error_general".Machine[1].Air_dryer;
         S     "DB009_Faults".Faultschanging_M1;

   // Fault air dryer --
   //    UN    "F_Airdryer_M2"
   //    UN    "DB820_Error_general".Machine[2].Air_dryer
   //    S     "DB820_Error_general".Machine[2].Air_dryer
   //    S     "DB009_Faults".Faultschanging_M2

   // Fault air dryer -- DB810.DBX 64.4
   //    UN    "P_SupplyAir"
   //    UN    "DB820_Error_general".Machine[1].P_AirSupply
   //    S     "DB820_Error_general".Machine[1].P_AirSupply
   //    S     "DB009_Faults".Faultschanging_M1

   // Fault heating general -- DB810.DBX 65.0
   //    UN    "F_SupplyHeatingM1"
   //    UN    "DB820_Error_general".Machine[1].Heating
   //    S     "DB820_Error_general".Machine[1].Heating
   //    S     "DB009_Faults".Faultschanging_M1

   // Fault pre alrarm Pentan  -- DB810.DBX 76.5
   //    UN    "K_PreAlarmN2_K1"
   //    UN    "DB820_Error_general".Machine[1].FLT_pre_alarm_pentan
   //    S     "DB820_Error_general".Machine[1].FLT_pre_alarm_pentan
   //    S     "DB009_Faults".Faultschanging_M1

   // Fault SGM faulty -- DB810.DBX 65.1
   //    UN      "K_SGM_Faulty"
   //    UN      "DB820_Error_general".Machine[1].SGM_Faulty
   //    S       "DB820_Error_general".Machine[1].SGM_Faulty
   //    S       "DB009_Faults".Faultschanging_M1

   // Automatic missing SGM -- DB810.DBX 65.6
   //    U       "DB123_MH_IO_Signals".MH[1].IN.MH_Auto_Mode
   //    U       "DB619_State_MPart".Operationmode_Ma[1].Auto
   //    UN      "K_SGM_Automatic"
   //    UN      "DB820_Error_general".Machine[1].SGM_AutomatcMissing
   //    S       "DB820_Error_general".Machine[1].SGM_AutomatcMissing
   //    S       "DB009_Faults".Faultschanging_M1

   // Fault Plasma  -- DB810.DBX 65.4
   //    UN    "K_PlasmaFaulty"
   //    UN    "DB820_Error_general".Machine[1].PlasmaFaulty
   //    S     "DB820_Error_general".Machine[1].PlasmaFaulty
   //    S     "DB009_Faults".Faultschanging_M1

   // Fault data transfer between PLC-memory and MMC -- DB810.DBX 77.5

   // Fault compressor cooling device -- DB810.DBX 65.2

         AN    "F_CoolingDevice";
         AN    "DB820_Error_general".Machine[1].F_CoolingDevice;
         S     "DB820_Error_general".Machine[1].F_CoolingDevice;
         S     "DB009_Faults".Faultschanging_M1;

   // Faults level 3 from PUC08
   //    U     "DB009_Faults".FaultPC_Level_3
   //    UN    "DB820_Error_general".Machine[1].FaultPC_Level_3
   //    S     "DB820_Error_general".Machine[1].FaultPC_Level_3
   //    S     "DB009_Faults".Faultschanging_M1

   //    U     "DB009_Faults".FaultPC_Level_3
   //    UN    "DB820_Error_general".Machine[2].FaultPC_Level_3
   //    S     "DB820_Error_general".Machine[2].FaultPC_Level_3
   //    S     "DB009_Faults".Faultschanging_M2

   //    O     "DB820_Error_general".Machine[1].FaultPC_Level_3
   //    O     "DB820_Error_general".Machine[1].Interface_PC
   //    O     "DB820_Error_general".Machine[1].BufferBattery
         O     "DB820_Error_general".Machine[1].Fuse_broken;
         O     "DB820_Error_general".Machine[1].Fuse_brocken_Mixinghead;
         O     "DB820_Error_general".Machine[1].Air_dryer;
         O     "DB820_Error_general".Machine[1].FLT_pre_alarm_pentan;
         O     "DB820_Error_general".Machine[1].SGM_Faulty;
         O     "DB820_Error_general".Machine[1].SGM_AutomatcMissing;
   //    O     "DB820_Error_general".Machine[1].TransferFaultMMC
         S     "DB009_Faults".Faults_FKT_Grp_3_M1;

   //    O     "DB820_Error_general".Machine[2].FaultPC_Level_3
   //    O     "DB820_Error_general".Machine[2].Interface_PC
   //    O     "DB820_Error_general".Machine[2].BufferBattery
         O     "DB820_Error_general".Machine[2].Fuse_broken;
         O     "DB820_Error_general".Machine[2].Fuse_brocken_Mixinghead;
         O     "DB820_Error_general".Machine[2].Air_dryer;
         O     "DB820_Error_general".Machine[2].FLT_pre_alarm_pentan;
         O     "DB820_Error_general".Machine[2].SGM_Faulty;
         O     "DB820_Error_general".Machine[2].SGM_AutomatcMissing;
   //    O     "DB820_Error_general".Machine[2].TransferFaultMMC
         S     "DB009_Faults".Faults_FKT_Grp_3_M2;
END_REGION

REGION Network 5: Messages

   // Controlvoltage maschine 1 missing  -- DB810.DBX64.5
   //-----------------------------------------------------------
         AN    "Controlvoltage";
         =     "DB820_Error_general".Machine[1].Controlvoltage;

   // Controlvoltage maschine 2 missing  --
   //-----------------------------------------------------------
   //    UN    "Controlvoltage_M2"
   //    =     "DB820_Error_general".Machine[2].Controlvoltage

   // Draining tank machine 1 -- DB810.DBX65.5
   //-----------------------------------------------------------
         O     "DB702_Tank_Value".Tank[1].DrainTank;
         O     "DB702_Tank_Value".Tank[2].DrainTank;
         O     "DB702_Tank_Value".Tank[3].DrainTank;
         O     "DB702_Tank_Value".Tank[4].DrainTank;
         =     "DB820_Error_general".Machine[1].DrainingTank;

   // Draining tank machine 2 -- DB810.DBX65.5
   //-----------------------------------------------------------
   //    O     "DB702_Tank_Refilling".Tank[3].DrainTank
   //    O     "DB702_Tank_Refilling".Tank[4].DrainTank
   //    =     "DB820_Error_general".Machine[2].DrainingTank

   // Not- Aus Taster an der Maschine wurde betätigt -- DB810.DBX66.0
   //------------------------------------------------------------
         A     "ES_Machine";
         =     "DB820_Error_general".Machine[1].EmergencyStop.Machine;

   // Not- Aus Taster an der Maschine wurde betätigt -- DB810.DBX66.0
   //    U     "ES_Machine_M2"
   //    =     "DB820_Error_general".Machine[2].EmergencyStop.Machine


   // Not- Aus Taster am Schaltschrank wurde betätigt -- DB810.DBX66.1
   //    =     "DB820_Error_general".EmergencyStop.Switch_Cabinet

   // Not- Aus Taster an dem Bedienpult der PUC08 wurde betätigt -- DB810.DBX66.2
   //-----------------------------------------------------------------------------
         A     "ES_Operatingpanel";
         =     "DB820_Error_general".Machine[1].EmergencyStop.Operation_Panel;

   // Not- Aus Taster am 2. Monitor wurde betätigt -- DB810.DBX66.3
   //    =      "DB820_Error_general".Machine[1].EmergencyStop.Monitor_2

   // Not- Aus Signal vom Roboter 1 steht an -- DB810.DBX66.7
         AN    "ES_Robot_01";
         CLR;
         =     "DB820_Error_general".Machine[1].EmergencyStop.Roboter_1;

   // Not- Aus Signal vom Roboter 2 steht an  -- DB810.DBX67.0
   //    UN    "ES_robot_MH2"
   //    =     "DB820_Error_general".Machine[2].EmergencyStop.Roboter_2

   // Not- Aus Taster an dem Behältern wurde betätigt
   //    =     "DB820_Error_general".Machine[1].EmergencyStop.Tank

   // Not- Aus Taster an dem Mischkopfreiniger 1 wurde betätigt -- DB810.DBX66.5
   //    =      "DB820_Error_general".Machine[1].EmergencyStop.MH_Cleaner_1

   // Not- Aus Taster an dem Mischkopfreiniger 2 wurde betätigt -- DB810.DBX66.6
         A     "ES_GBE_C1";
         A     "DB702_Tank_Value".Tank[1].With_Nucleation;
         =     "DB820_Error_general".Machine[1].EmergencyStop.MH_Cleaner_2;